(* Logix 5000 project; controller _GigaDiscovery vendor 1 type 14 code 244 rev 35.11; software revision 35.03; part 22 of 23 *)
(* tags used below, declared in another part *)
   All_Rack_Closed_Mem : BOOL;
   Close_Platform_Autocycle_Pylon : BOOL;
   CycleOver : BOOL;
   Emergencies_CL0 : DINT[8];
   FeedBack_Drives_Contactors : BOOL;
   GateCommand : DINT;
   GateRequest : DINT;
   Gates_Auto_Release : BOOL;   // .. At end of Cycle Open Gates Open RESTRAINTS
   Gates_Open_Permissive : Permissive;
   Gondola_Standstill_from_inertia : BOOL;
   HMI_PAGE_PROOF_TEST : DINT;
   I_EStop_Pb_OCC1 : UDT_DCI_STOP_TEST;   // +OCC E-stop -S30301F
   I_EStop_Pb_OCC2 : UDT_DCI_STOP_TEST;   // +OCC2 E-Stop -S28502F
   I_Gondola_Home_Position : BOOL;   // Gondola Home Position -B40002I -B40007I
   I_OCC1_EntGate_PB : BOOL;   // OCC1 Entrance Gate Open/Close -S30701F
   I_OCC1_ExitGate_PB : BOOL;   // OCC1 ExitGate Open/Close -S30707F
   I_OCC2_Disable : UDT_DCM;   // OCC 2 CONTROL DISABLE Page 310
   I_OCC2_ExitGate_PB : BOOL;   // OCC2 ExitGate Open/Close -S28507F
   I_OCC2_RESTRAINTS_RELEASE : Sel_3_Pos_2_Input;   // -S28507F RESTRAINTS RELEASE UNLOCK -RUN- LOCK
   I_OCC_LockOut_Motion : UDT_DCM;   // OCC -Lockout Motion -Q31203E
   I_OCC_Operator_Enable_Key : BOOL;   // OCC Console Enabled -S30305F
   I_Platform_Closed : UDT_DCM;   // Platform Closed RFID Series -B22501J... -B22807J -B22801B
   I_Platform_Line_Min_Pressure_Switch : BOOL;   // Platform Line Minimum Pressure Switch -S21511B
   I_Platform_Line_Unlock_Pressure_Switch : BOOL;   // Unlock Platform Line Pressure Switch -S22006B
   I_Platform_Pressure_on_Close_Circuit : BOOL;   // Platform Maximum Closing Pressure -S21510B
   I_RESTRAINTS_Selector : Sel_3_Pos_2_Input;   // RESTRAINTS Selctor -S30505F Left = Open Right = Close Center = Nothing
   Mem_RESTRAINTS_closed_Correctly : BOOL;
   No_Sfty : Std_to_Sfty;
   O_Close_Gate1 : BOOL;   // Gate 1 OCC2 Operator Close = Mag ON
   O_Close_Gate2 : BOOL;   // Gate 2 Exit Close = Mag ON
   O_Close_Gate3 : BOOL;   // Gate 3 Entrance Close = Mag ON
   O_Close_Gates : BOOL;
   O_Close_Platform : BOOL;
   O_Open_Platform : BOOL;
   O_Platform_Main_Valve : BOOL;   // Valvola principale piattaforma B21902I
   O_RESTRAINTS_MainValve : UDT_CROUT;   // Main Valve -B40501I
   O_RESTRAINTS_Valve_Lift : BOOL;   // Steps 03 04 05
   OS_Start_Stop_Cycle_Started : BOOL;
   Paltform_Cycle_Abborted_Mem : BOOL;   // Paltform Cycle Abborted by Stop Pb Mem
   Pb_Platform_Stop : BOOL;   // Platform Stop Command -S30608F
   PltaformClosed_CycleComplete : BOOL;   // Piattaforme chiuse e ciclo completato
   Power_On_Delay : BOOL;
   ProofTest_Req : BOOL;
   Pylon_Contactor_OFF : BOOL;
   Pylon_Stopped_At_Home : BOOL;   // 5s
   RESTRAINTS_Closed : BOOL;   // All RESTRAINTS Closed
   Restraints_Cycle : Sequencer;
   RESTRAINTS_Left_Press_Switch_Series : BOOL;
   RESTRAINTS_No_Alarms : BOOL;
   Restraints_Permissive : Permissive;
   Restraints_Permissive_Ok : BOOL;
   Restraints_PermissiveLost : DINT;
   RESTRAINTS_Right_Press_Switch_Series : BOOL;
   RESTRAINTS_Sector : LapBars_Sector[9];
   Start_Stop_Cycle : Sequencer;
   Test : DCI_STOP_TEST;
(* S_Platform_and_Gates, continued *)

ROUTINE _10_Gates_Permissive   (* ladder *)
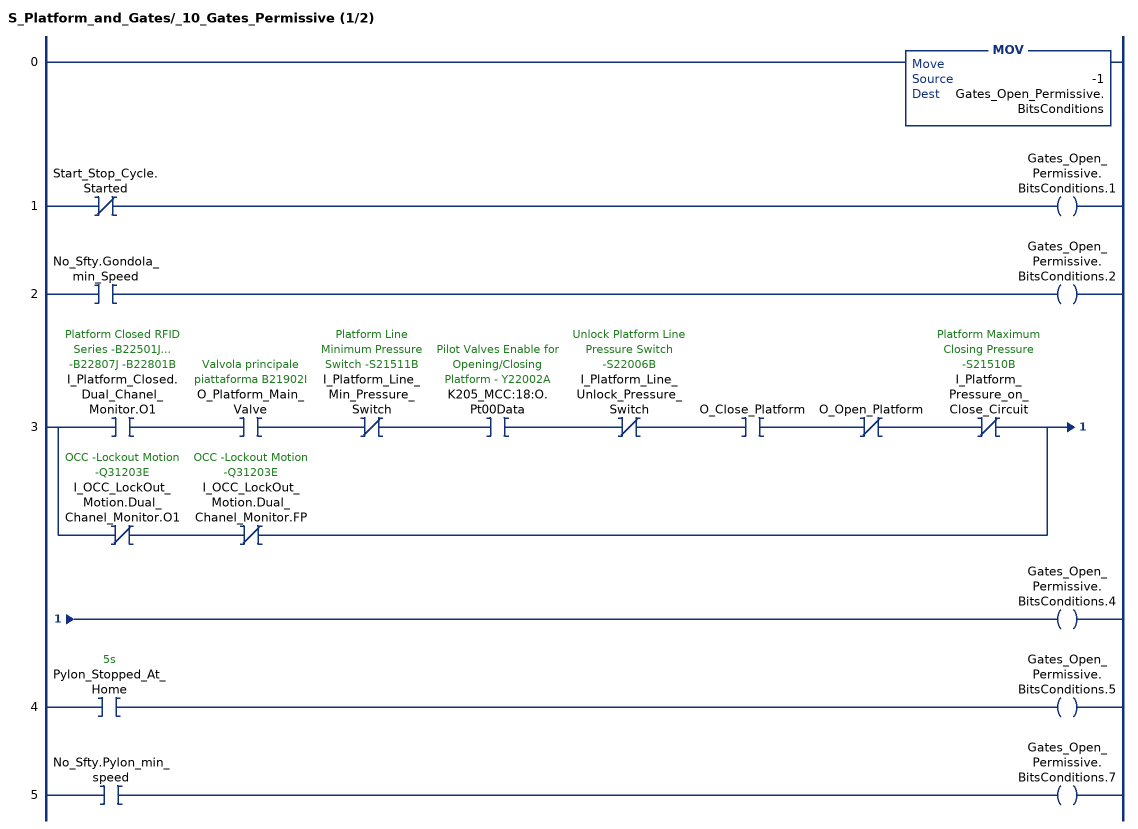
   0: MOV(-1,Gates_Open_Permissive.BitsConditions);
   1: XIO(Start_Stop_Cycle.Started)OTE(Gates_Open_Permissive.BitsConditions.1);
   2: XIC(No_Sfty.Gondola_min_Speed)OTE(Gates_Open_Permissive.BitsConditions.2);
   3: [XIC(I_Platform_Closed.Dual_Chanel_Monitor.O1) XIC(O_Platform_Main_Valve) XIO(I_Platform_Line_Min_Pressure_Switch) XIC(K205_MCC:18:O.Pt00Data) XIO(I_Platform_Line_Unlock_Pressure_Switch) XIC(O_Close_Platform) XIO(O_Open_Platform) XIO(I_Platform_Pressure_on_Close_Circuit) ,XIO(I_OCC_LockOut_Motion.Dual_Chanel_Monitor.O1) XIO(I_OCC_LockOut_Motion.Dual_Chanel_Monitor.FP) ]OTE(Gates_Open_Permissive.BitsConditions.4);
   4: XIC(Pylon_Stopped_At_Home)OTE(Gates_Open_Permissive.BitsConditions.5);
   5: XIC(No_Sfty.Pylon_min_speed)OTE(Gates_Open_Permissive.BitsConditions.7);
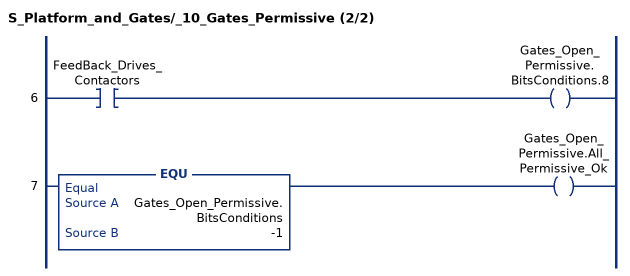
   6: XIC(FeedBack_Drives_Contactors)OTE(Gates_Open_Permissive.BitsConditions.8);
   7: EQU(Gates_Open_Permissive.BitsConditions,-1)OTE(Gates_Open_Permissive.All_Permissive_Ok);
END_ROUTINE

ROUTINE _11_Gates_Commands   (* ladder *)
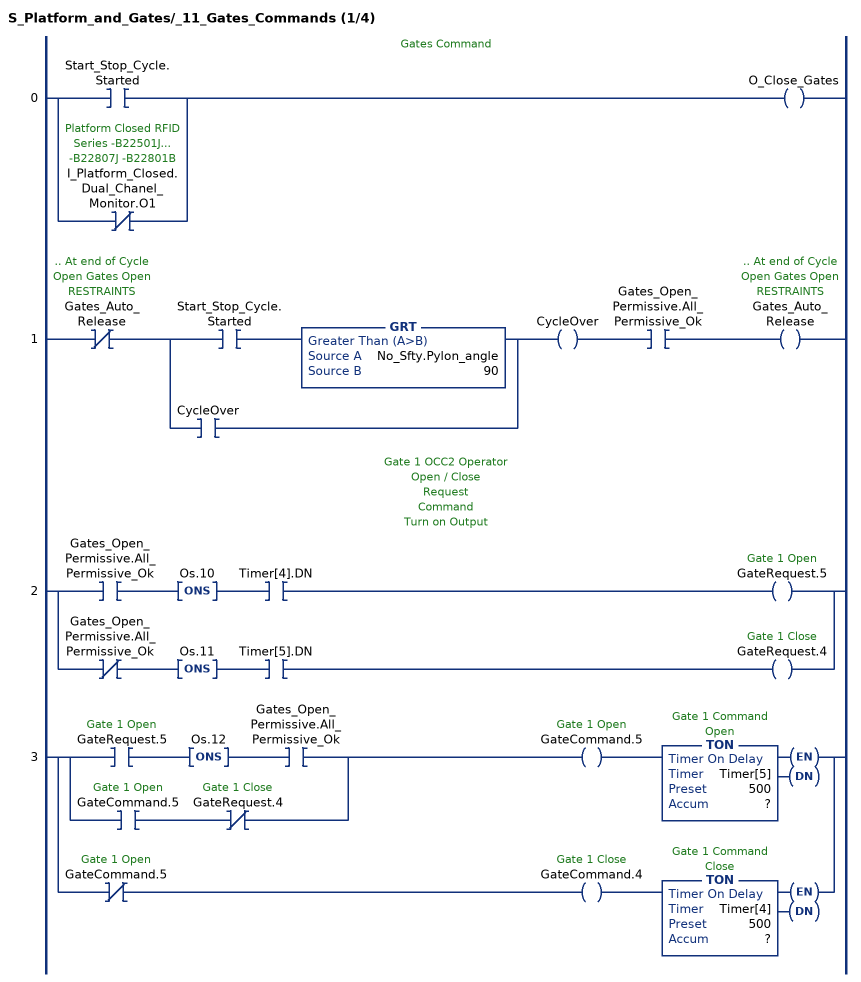
   // Gates Command
   0: [XIC(Start_Stop_Cycle.Started) ,XIO(I_Platform_Closed.Dual_Chanel_Monitor.O1) ]OTE(O_Close_Gates);
   1: XIO(Gates_Auto_Release)[XIC(Start_Stop_Cycle.Started) GRT(No_Sfty.Pylon_angle,90) ,XIC(CycleOver) ]OTE(CycleOver)XIC(Gates_Open_Permissive.All_Permissive_Ok)OTE(Gates_Auto_Release);
   // Gate 1 OCC2 Operator
   // Open / Close
   // Request
   // Command
   // Turn on Output
   2: [XIC(Gates_Open_Permissive.All_Permissive_Ok) ONS(Os.10) XIC(Timer[4].DN) OTE(GateRequest.5) ,XIO(Gates_Open_Permissive.All_Permissive_Ok) ONS(Os.11) XIC(Timer[5].DN) OTE(GateRequest.4) ];
   3: [[XIC(GateRequest.5) ONS(Os.12) XIC(Gates_Open_Permissive.All_Permissive_Ok) ,XIC(GateCommand.5) XIO(GateRequest.4) ] OTE(GateCommand.5) TON(Timer[5],?,?) ,XIO(GateCommand.5) OTE(GateCommand.4) TON(Timer[4],?,?) ];
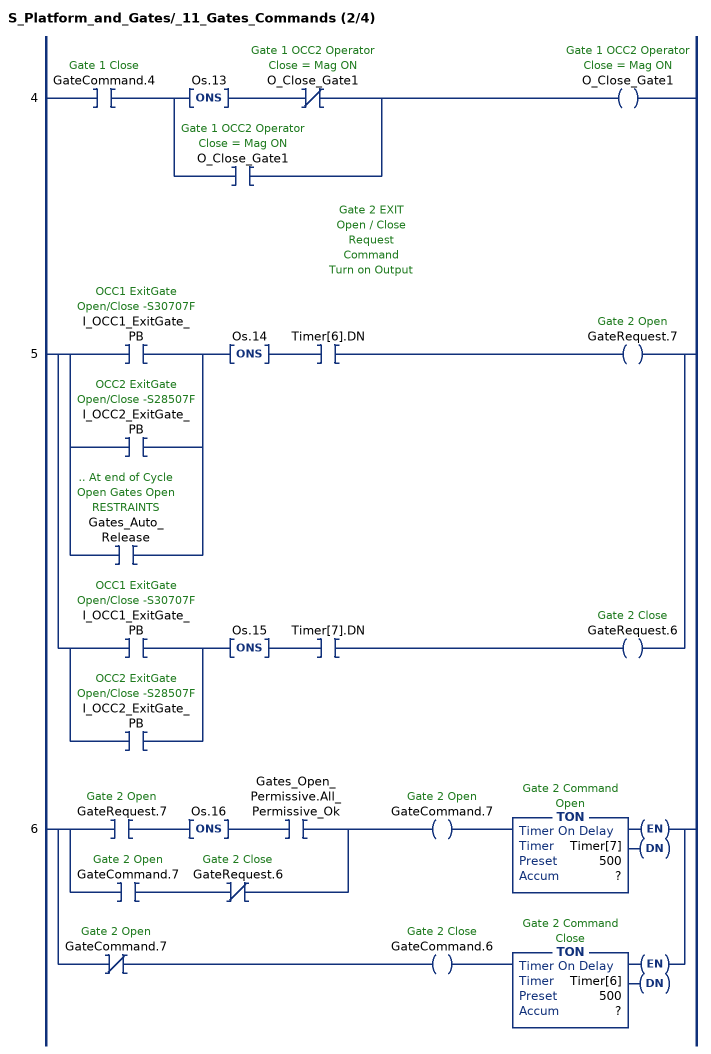
   4: XIC(GateCommand.4)[ONS(Os.13) XIO(O_Close_Gate1) ,XIC(O_Close_Gate1) ]OTE(O_Close_Gate1);
   // Gate 2 EXIT
   // Open / Close
   // Request
   // Command
   // Turn on Output
   5: [[XIC(I_OCC1_ExitGate_PB) ,XIC(I_OCC2_ExitGate_PB) ,XIC(Gates_Auto_Release) ] ONS(Os.14) XIC(Timer[6].DN) OTE(GateRequest.7) ,[XIC(I_OCC1_ExitGate_PB) ,XIC(I_OCC2_ExitGate_PB) ] ONS(Os.15) XIC(Timer[7].DN) OTE(GateRequest.6) ];
   6: [[XIC(GateRequest.7) ONS(Os.16) XIC(Gates_Open_Permissive.All_Permissive_Ok) ,XIC(GateCommand.7) XIO(GateRequest.6) ] OTE(GateCommand.7) TON(Timer[7],?,?) ,XIO(GateCommand.7) OTE(GateCommand.6) TON(Timer[6],?,?) ];
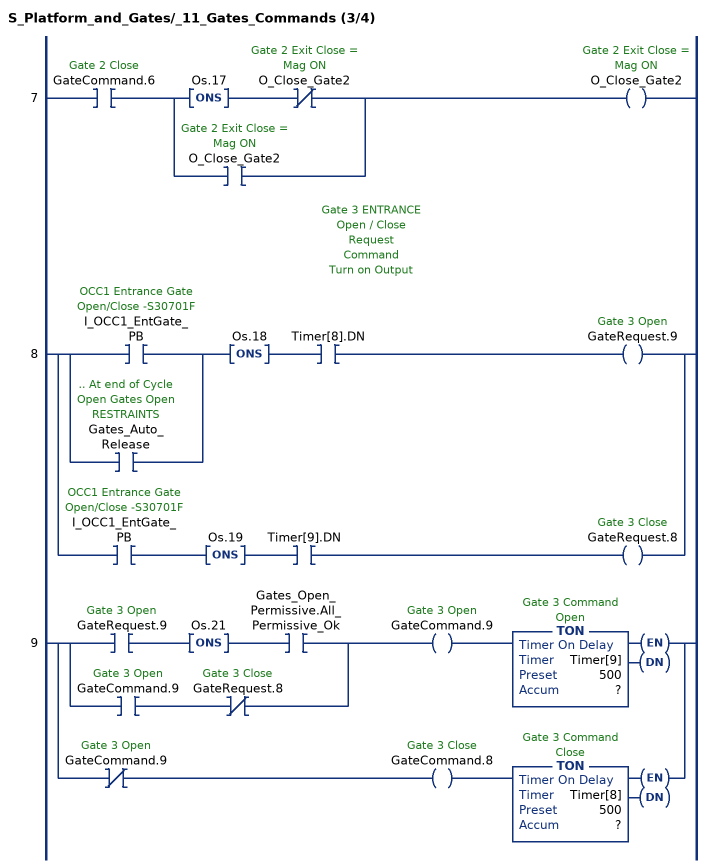
   7: XIC(GateCommand.6)[ONS(Os.17) XIO(O_Close_Gate2) ,XIC(O_Close_Gate2) ]OTE(O_Close_Gate2);
   // Gate 3 ENTRANCE
   // Open / Close
   // Request
   // Command
   // Turn on Output
   8: [[XIC(I_OCC1_EntGate_PB) ,XIC(Gates_Auto_Release) ] ONS(Os.18) XIC(Timer[8].DN) OTE(GateRequest.9) ,XIC(I_OCC1_EntGate_PB) ONS(Os.19) XIC(Timer[9].DN) OTE(GateRequest.8) ];
   9: [[XIC(GateRequest.9) ONS(Os.21) XIC(Gates_Open_Permissive.All_Permissive_Ok) ,XIC(GateCommand.9) XIO(GateRequest.8) ] OTE(GateCommand.9) TON(Timer[9],?,?) ,XIO(GateCommand.9) OTE(GateCommand.8) TON(Timer[8],?,?) ];
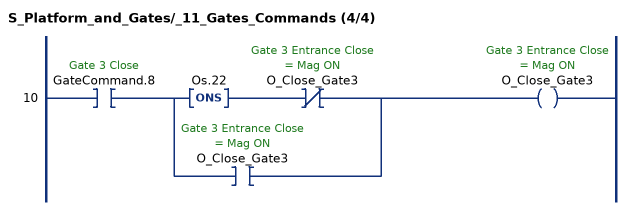
   10: XIC(GateCommand.8)[ONS(Os.22) XIO(O_Close_Gate3) ,XIC(O_Close_Gate3) ]OTE(O_Close_Gate3);
END_ROUTINE

ROUTINE Main   (* ladder *)
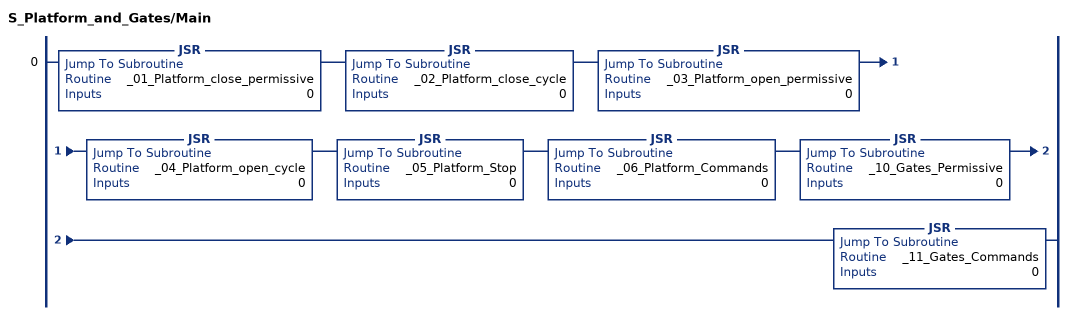
   0: JSR(_01_Platform_close_permissive,0)JSR(_02_Platform_close_cycle,0)JSR(_03_Platform_open_permissive,0)JSR(_04_Platform_open_cycle,0)JSR(_05_Platform_Stop,0)JSR(_06_Platform_Commands,0)JSR(_10_Gates_Permissive,0)JSR(_11_Gates_Commands,0);
END_ROUTINE
END_PROGRAM

PROGRAM S_Restraints_Release   (* main routine Main, safety *)
VAR
   _07_Stop_RESTRAINT_RELEASE_Cycle : BOOL;
   O_Safety_Valve_Unlock_Left_Block : BOOL;   // Steps 02 to 21
   O_Safety_Valve_Unlock_Right_Block : BOOL;   // Steps 02 to 21
   Os : DINT := 45040;
   Proof_Test : Proof_Test := (Validation_Delay_time.PRE := 30000);
   Proof_Test_Req_by_Time : BOOL;
   RESTRAINT_RELEASE_Alarm_Loc : BOOL;
   RESTRAINT_RELEASE_Cycle_AOI : Sequencer_AOI;
   Timer : TIMER[11] := ([0].PRE := 60000, [1].PRE := 2000, [1].ACC := 2000, [1].EN := 1, [1].DN := 1);
END_VAR

ROUTINE _01_Restraints_Release_Permissives   (* ladder *)
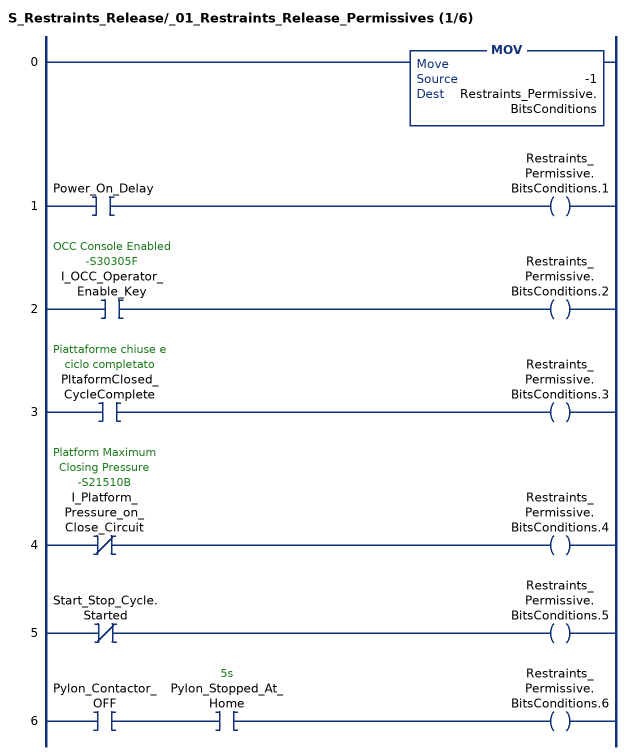
   0: MOV(-1,Restraints_Permissive.BitsConditions);
   1: XIC(Power_On_Delay)OTE(Restraints_Permissive.BitsConditions.1);
   2: XIC(I_OCC_Operator_Enable_Key)OTE(Restraints_Permissive.BitsConditions.2);
   3: XIC(PltaformClosed_CycleComplete)OTE(Restraints_Permissive.BitsConditions.3);
   4: XIO(I_Platform_Pressure_on_Close_Circuit)OTE(Restraints_Permissive.BitsConditions.4);
   5: XIO(Start_Stop_Cycle.Started)OTE(Restraints_Permissive.BitsConditions.5);
   6: XIC(Pylon_Contactor_OFF)XIC(Pylon_Stopped_At_Home)OTE(Restraints_Permissive.BitsConditions.6);
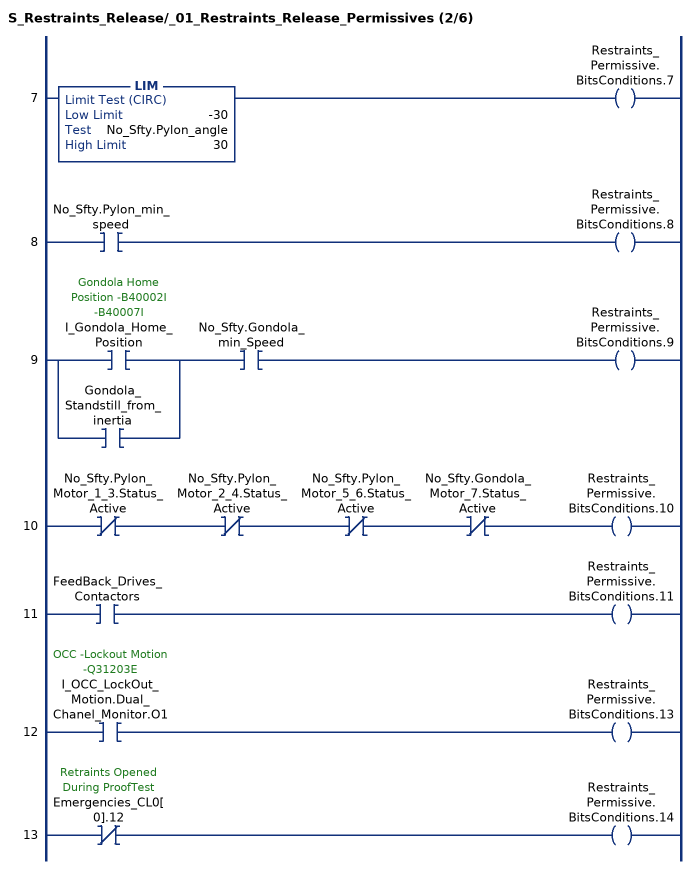
   7: LIM(-30,No_Sfty.Pylon_angle,30)OTE(Restraints_Permissive.BitsConditions.7);
   8: XIC(No_Sfty.Pylon_min_speed)OTE(Restraints_Permissive.BitsConditions.8);
   9: [XIC(I_Gondola_Home_Position) ,XIC(Gondola_Standstill_from_inertia) ]XIC(No_Sfty.Gondola_min_Speed)OTE(Restraints_Permissive.BitsConditions.9);
   10: XIO(No_Sfty.Pylon_Motor_1_3.Status_Active)XIO(No_Sfty.Pylon_Motor_2_4.Status_Active)XIO(No_Sfty.Pylon_Motor_5_6.Status_Active)XIO(No_Sfty.Gondola_Motor_7.Status_Active)OTE(Restraints_Permissive.BitsConditions.10);
   11: XIC(FeedBack_Drives_Contactors)OTE(Restraints_Permissive.BitsConditions.11);
   12: XIC(I_OCC_LockOut_Motion.Dual_Chanel_Monitor.O1)OTE(Restraints_Permissive.BitsConditions.13);
   13: XIO(Emergencies_CL0[0].12)OTE(Restraints_Permissive.BitsConditions.14);
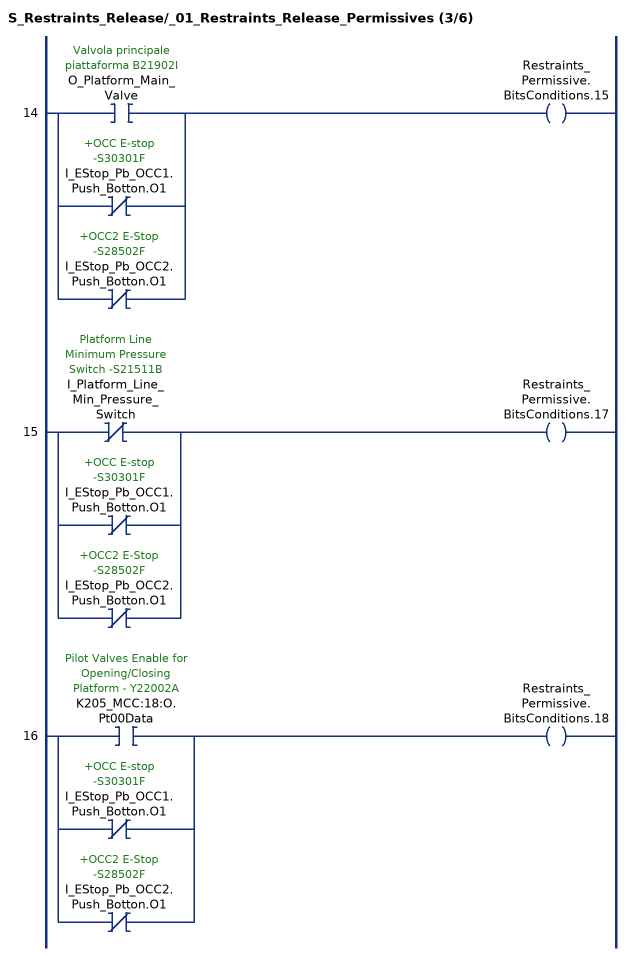
   14: [XIC(O_Platform_Main_Valve) ,XIO(I_EStop_Pb_OCC1.Push_Botton.O1) ,XIO(I_EStop_Pb_OCC2.Push_Botton.O1) ]OTE(Restraints_Permissive.BitsConditions.15);
   15: [XIO(I_Platform_Line_Min_Pressure_Switch) ,XIO(I_EStop_Pb_OCC1.Push_Botton.O1) ,XIO(I_EStop_Pb_OCC2.Push_Botton.O1) ]OTE(Restraints_Permissive.BitsConditions.17);
   16: [XIC(K205_MCC:18:O.Pt00Data) ,XIO(I_EStop_Pb_OCC1.Push_Botton.O1) ,XIO(I_EStop_Pb_OCC2.Push_Botton.O1) ]OTE(Restraints_Permissive.BitsConditions.18);
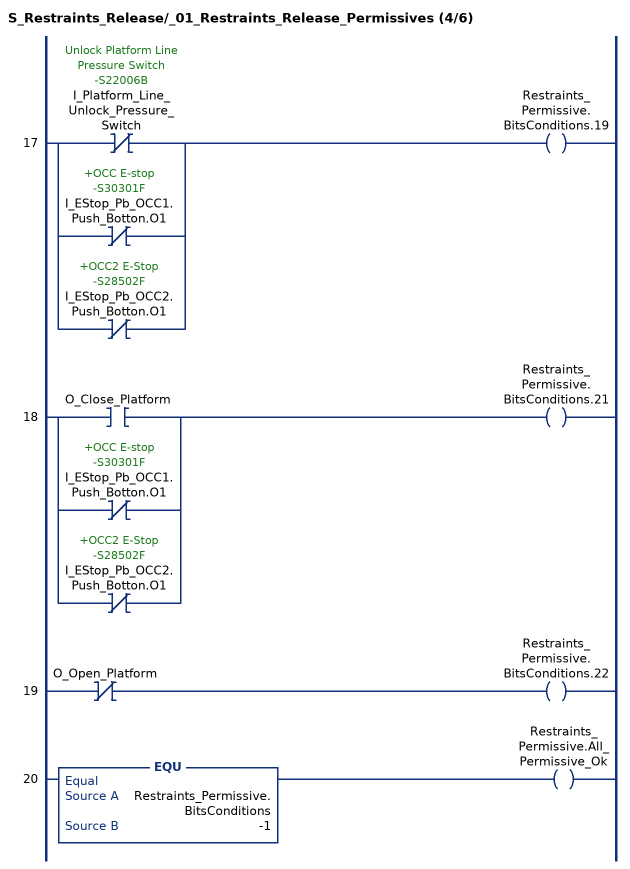
   17: [XIO(I_Platform_Line_Unlock_Pressure_Switch) ,XIO(I_EStop_Pb_OCC1.Push_Botton.O1) ,XIO(I_EStop_Pb_OCC2.Push_Botton.O1) ]OTE(Restraints_Permissive.BitsConditions.19);
   18: [XIC(O_Close_Platform) ,XIO(I_EStop_Pb_OCC1.Push_Botton.O1) ,XIO(I_EStop_Pb_OCC2.Push_Botton.O1) ]OTE(Restraints_Permissive.BitsConditions.21);
   19: XIO(O_Open_Platform)OTE(Restraints_Permissive.BitsConditions.22);
   20: EQU(Restraints_Permissive.BitsConditions,-1)OTE(Restraints_Permissive.All_Permissive_Ok);
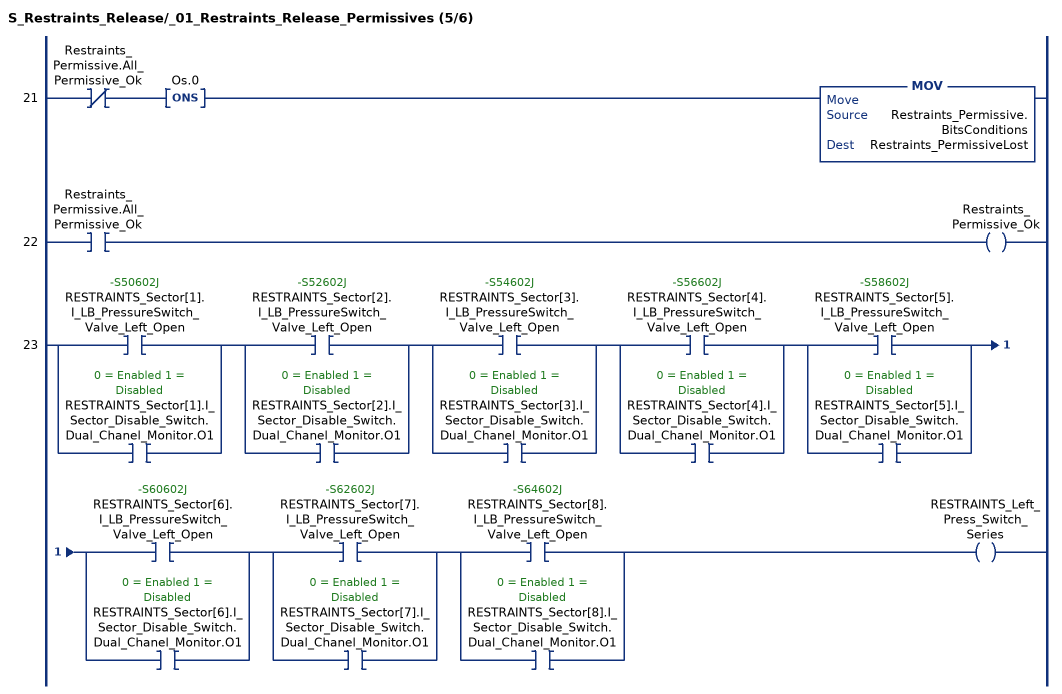
   21: XIO(Restraints_Permissive.All_Permissive_Ok)ONS(Os.0)MOV(Restraints_Permissive.BitsConditions,Restraints_PermissiveLost);
   22: XIC(Restraints_Permissive.All_Permissive_Ok)OTE(Restraints_Permissive_Ok);
   23: [XIC(RESTRAINTS_Sector[1].I_LB_PressureSwitch_Valve_Left_Open) ,XIC(RESTRAINTS_Sector[1].I_Sector_Disable_Switch.Dual_Chanel_Monitor.O1) ][XIC(RESTRAINTS_Sector[2].I_LB_PressureSwitch_Valve_Left_Open) ,XIC(RESTRAINTS_Sector[2].I_Sector_Disable_Switch.Dual_Chanel_Monitor.O1) ][XIC(RESTRAINTS_Sector[3].I_LB_PressureSwitch_Valve_Left_Open) ,XIC(RESTRAINTS_Sector[3].I_Sector_Disable_Switch.Dual_Chanel_Monitor.O1) ][XIC(RESTRAINTS_Sector[4].I_LB_PressureSwitch_Valve_Left_Open) ,XIC(RESTRAINTS_Sector[4].I_Sector_Disable_Switch.Dual_Chanel_Monitor.O1) ][XIC(RESTRAINTS_Sector[5].I_LB_PressureSwitch_Valve_Left_Open) ,XIC(RESTRAINTS_Sector[5].I_Sector_Disable_Switch.Dual_Chanel_Monitor.O1) ][XIC(RESTRAINTS_Sector[6].I_LB_PressureSwitch_Valve_Left_Open) ,XIC(RESTRAINTS_Sector[6].I_Sector_Disable_Switch.Dual_Chanel_Monitor.O1) ][XIC(RESTRAINTS_Sector[7].I_LB_PressureSwitch_Valve_Left_Open) ,XIC(RESTRAINTS_Sector[7].I_Sector_Disable_Switch.Dual_Chanel_Monitor.O1) ][XIC(RESTRAINTS_Sector[8].I_LB_PressureSwitch_Valve_Left_Open) ,XIC(RESTRAINTS_Sector[8].I_Sector_Disable_Switch.Dual_Chanel_Monitor.O1) ]OTE(RESTRAINTS_Left_Press_Switch_Series);
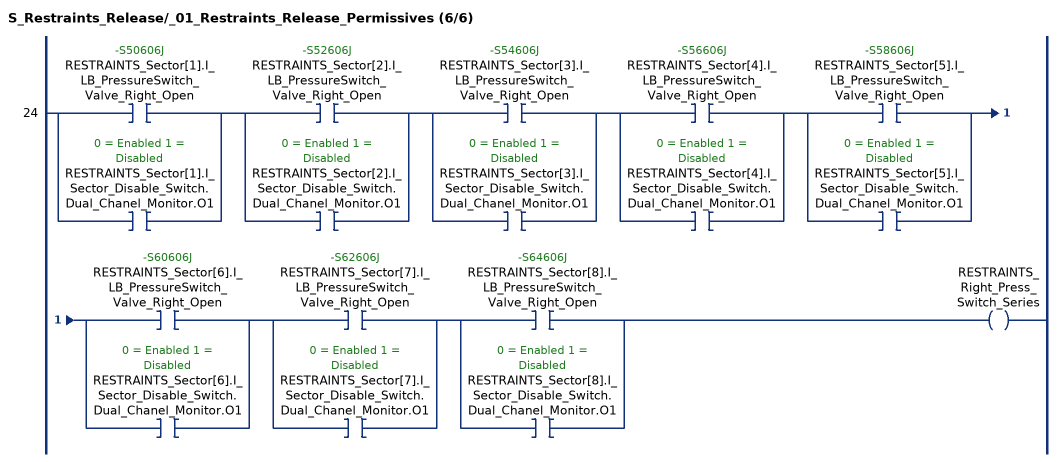
   24: [XIC(RESTRAINTS_Sector[1].I_LB_PressureSwitch_Valve_Right_Open) ,XIC(RESTRAINTS_Sector[1].I_Sector_Disable_Switch.Dual_Chanel_Monitor.O1) ][XIC(RESTRAINTS_Sector[2].I_LB_PressureSwitch_Valve_Right_Open) ,XIC(RESTRAINTS_Sector[2].I_Sector_Disable_Switch.Dual_Chanel_Monitor.O1) ][XIC(RESTRAINTS_Sector[3].I_LB_PressureSwitch_Valve_Right_Open) ,XIC(RESTRAINTS_Sector[3].I_Sector_Disable_Switch.Dual_Chanel_Monitor.O1) ][XIC(RESTRAINTS_Sector[4].I_LB_PressureSwitch_Valve_Right_Open) ,XIC(RESTRAINTS_Sector[4].I_Sector_Disable_Switch.Dual_Chanel_Monitor.O1) ][XIC(RESTRAINTS_Sector[5].I_LB_PressureSwitch_Valve_Right_Open) ,XIC(RESTRAINTS_Sector[5].I_Sector_Disable_Switch.Dual_Chanel_Monitor.O1) ][XIC(RESTRAINTS_Sector[6].I_LB_PressureSwitch_Valve_Right_Open) ,XIC(RESTRAINTS_Sector[6].I_Sector_Disable_Switch.Dual_Chanel_Monitor.O1) ][XIC(RESTRAINTS_Sector[7].I_LB_PressureSwitch_Valve_Right_Open) ,XIC(RESTRAINTS_Sector[7].I_Sector_Disable_Switch.Dual_Chanel_Monitor.O1) ][XIC(RESTRAINTS_Sector[8].I_LB_PressureSwitch_Valve_Right_Open) ,XIC(RESTRAINTS_Sector[8].I_Sector_Disable_Switch.Dual_Chanel_Monitor.O1) ]OTE(RESTRAINTS_Right_Press_Switch_Series);
END_ROUTINE

ROUTINE _02_Restraints_Release_Cycle   (* ladder *)
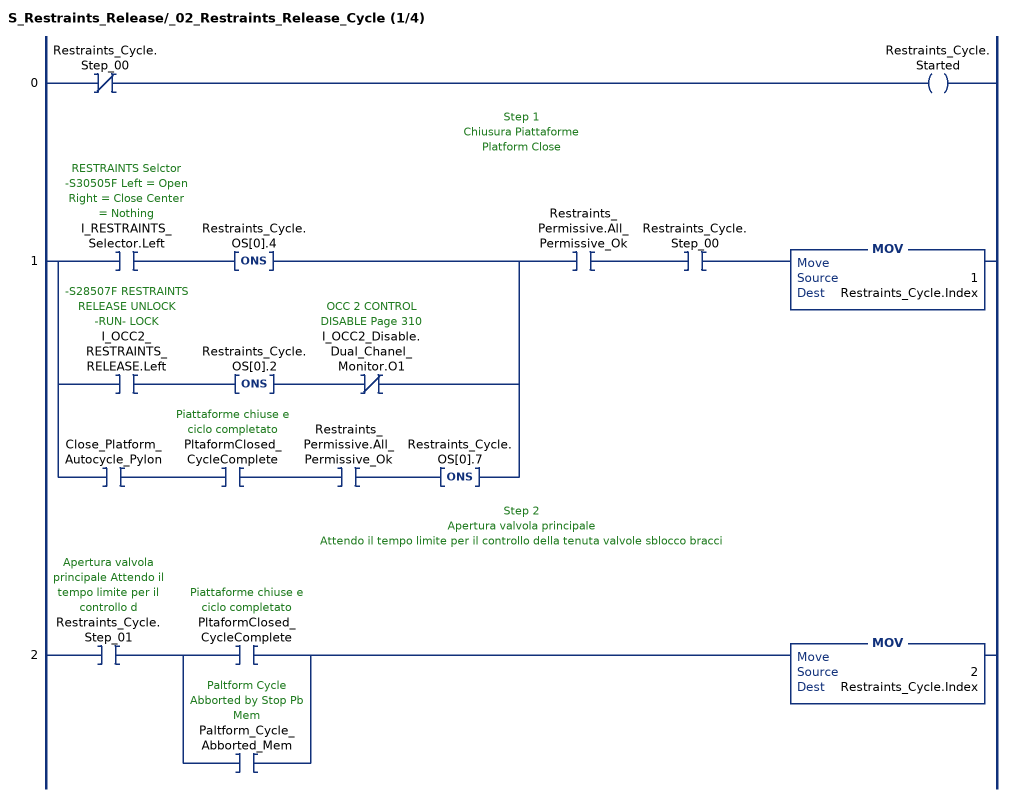
   0: XIO(Restraints_Cycle.Step_00)OTE(Restraints_Cycle.Started);
   // Step 1
   // Chiusura Piattaforme
   // Platform Close
   1: [XIC(I_RESTRAINTS_Selector.Left) ONS(Restraints_Cycle.OS[0].4) ,XIC(I_OCC2_RESTRAINTS_RELEASE.Left) ONS(Restraints_Cycle.OS[0].2) XIO(I_OCC2_Disable.Dual_Chanel_Monitor.O1) ,XIC(Close_Platform_Autocycle_Pylon) XIC(PltaformClosed_CycleComplete) XIC(Restraints_Permissive.All_Permissive_Ok) ONS(Restraints_Cycle.OS[0].7) ]XIC(Restraints_Permissive.All_Permissive_Ok)XIC(Restraints_Cycle.Step_00)MOV(1,Restraints_Cycle.Index);
   // Step 2
   // Apertura valvola principale
   // Attendo il tempo limite per il controllo della tenuta valvole sblocco bracci
   2: XIC(Restraints_Cycle.Step_01)[XIC(PltaformClosed_CycleComplete) ,XIC(Paltform_Cycle_Abborted_Mem) ]MOV(2,Restraints_Cycle.Index);
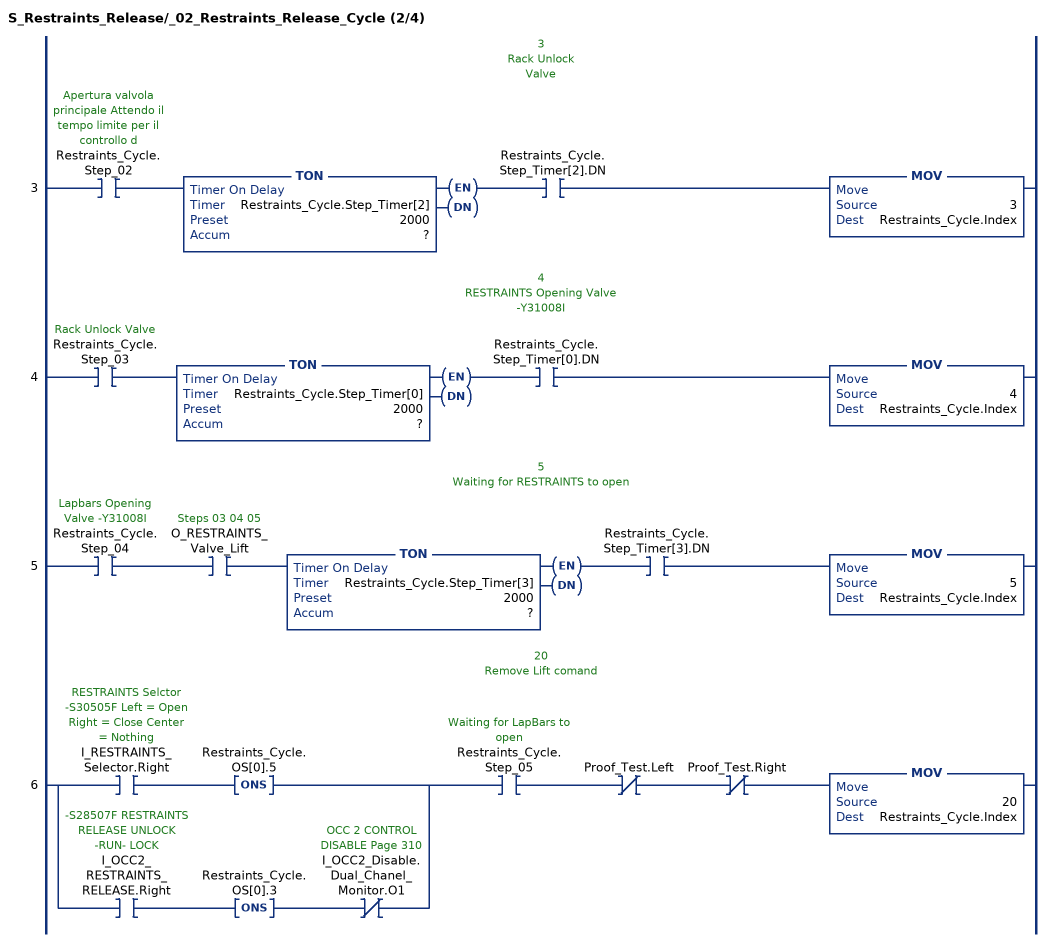
   // 3
   // Rack Unlock
   // Valve
   3: XIC(Restraints_Cycle.Step_02)TON(Restraints_Cycle.Step_Timer[2],?,?)XIC(Restraints_Cycle.Step_Timer[2].DN)MOV(3,Restraints_Cycle.Index);
   // 4
   // RESTRAINTS Opening Valve
   // -Y31008I
   4: XIC(Restraints_Cycle.Step_03)TON(Restraints_Cycle.Step_Timer[0],?,?)XIC(Restraints_Cycle.Step_Timer[0].DN)MOV(4,Restraints_Cycle.Index);
   // 5
   // Waiting for RESTRAINTS to open
   5: XIC(Restraints_Cycle.Step_04)XIC(O_RESTRAINTS_Valve_Lift)TON(Restraints_Cycle.Step_Timer[3],?,?)XIC(Restraints_Cycle.Step_Timer[3].DN)MOV(5,Restraints_Cycle.Index);
   // 20
   // Remove Lift comand
   6: [XIC(I_RESTRAINTS_Selector.Right) ONS(Restraints_Cycle.OS[0].5) ,XIC(I_OCC2_RESTRAINTS_RELEASE.Right) ONS(Restraints_Cycle.OS[0].3) XIO(I_OCC2_Disable.Dual_Chanel_Monitor.O1) ]XIC(Restraints_Cycle.Step_05)XIO(Proof_Test.Left)XIO(Proof_Test.Right)MOV(20,Restraints_Cycle.Index);
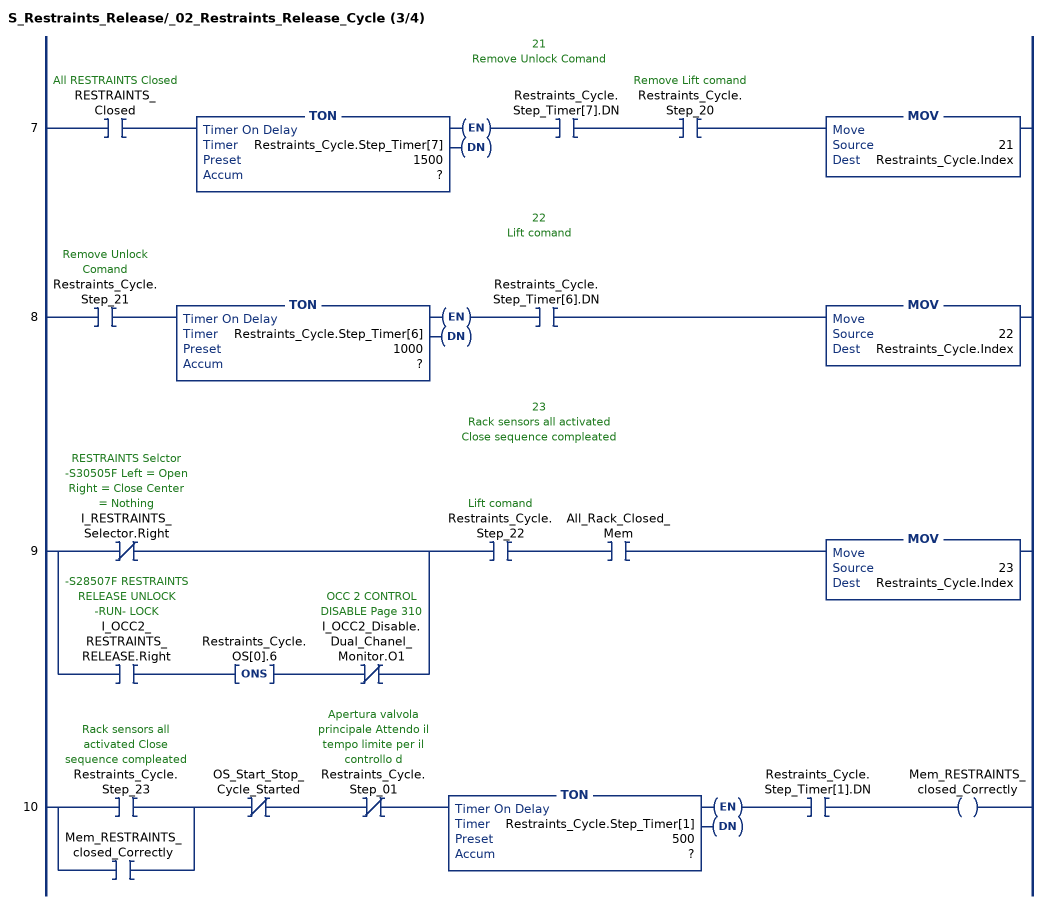
   // 21
   // Remove Unlock Comand
   7: XIC(RESTRAINTS_Closed)TON(Restraints_Cycle.Step_Timer[7],?,?)XIC(Restraints_Cycle.Step_Timer[7].DN)XIC(Restraints_Cycle.Step_20)MOV(21,Restraints_Cycle.Index);
   // 22
   // Lift comand
   8: XIC(Restraints_Cycle.Step_21)TON(Restraints_Cycle.Step_Timer[6],?,?)XIC(Restraints_Cycle.Step_Timer[6].DN)MOV(22,Restraints_Cycle.Index);
   // 23
   // Rack sensors all activated
   // Close sequence compleated
   9: [XIO(I_RESTRAINTS_Selector.Right) ,XIC(I_OCC2_RESTRAINTS_RELEASE.Right) ONS(Restraints_Cycle.OS[0].6) XIO(I_OCC2_Disable.Dual_Chanel_Monitor.O1) ]XIC(Restraints_Cycle.Step_22)XIC(All_Rack_Closed_Mem)MOV(23,Restraints_Cycle.Index);
   10: [XIC(Restraints_Cycle.Step_23) ,XIC(Mem_RESTRAINTS_closed_Correctly) ]XIO(OS_Start_Stop_Cycle_Started)XIO(Restraints_Cycle.Step_01)TON(Restraints_Cycle.Step_Timer[1],?,?)XIC(Restraints_Cycle.Step_Timer[1].DN)OTE(Mem_RESTRAINTS_closed_Correctly);
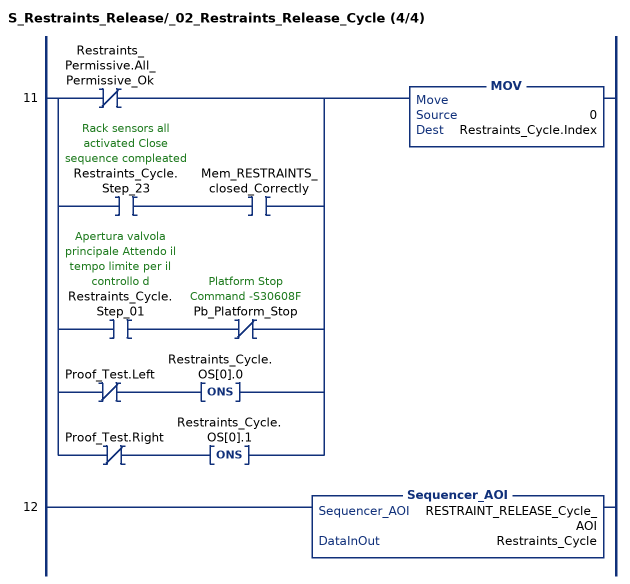
   11: [XIO(Restraints_Permissive.All_Permissive_Ok) ,XIC(Restraints_Cycle.Step_23) XIC(Mem_RESTRAINTS_closed_Correctly) ,XIC(Restraints_Cycle.Step_01) XIO(Pb_Platform_Stop) ,XIO(Proof_Test.Left) ONS(Restraints_Cycle.OS[0].0) ,XIO(Proof_Test.Right) ONS(Restraints_Cycle.OS[0].1) ]MOV(0,Restraints_Cycle.Index);
   12: Sequencer_AOI(RESTRAINT_RELEASE_Cycle_AOI,Restraints_Cycle);
END_ROUTINE

ROUTINE _03_Proof_Test   (* ladder *)
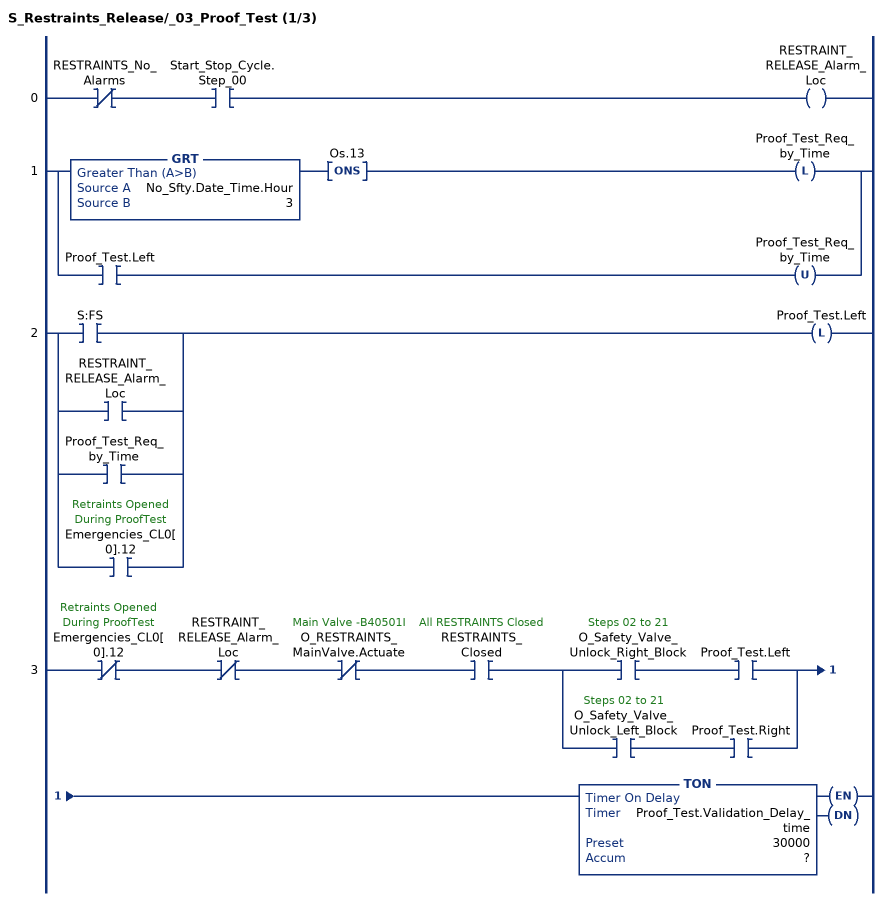
   0: XIO(RESTRAINTS_No_Alarms)XIC(Start_Stop_Cycle.Step_00)OTE(RESTRAINT_RELEASE_Alarm_Loc);
   1: [GRT(No_Sfty.Date_Time.Hour,3) ONS(Os.13) OTL(Proof_Test_Req_by_Time) ,XIC(Proof_Test.Left) OTU(Proof_Test_Req_by_Time) ];
   2: [XIC(S:FS) ,XIC(RESTRAINT_RELEASE_Alarm_Loc) ,XIC(Proof_Test_Req_by_Time) ,XIC(Emergencies_CL0[0].12) ]OTL(Proof_Test.Left);
   3: XIO(Emergencies_CL0[0].12)XIO(RESTRAINT_RELEASE_Alarm_Loc)XIO(O_RESTRAINTS_MainValve.Actuate)XIC(RESTRAINTS_Closed)[XIC(O_Safety_Valve_Unlock_Right_Block) XIC(Proof_Test.Left) ,XIC(O_Safety_Valve_Unlock_Left_Block) XIC(Proof_Test.Right) ]TON(Proof_Test.Validation_Delay_time,?,?);
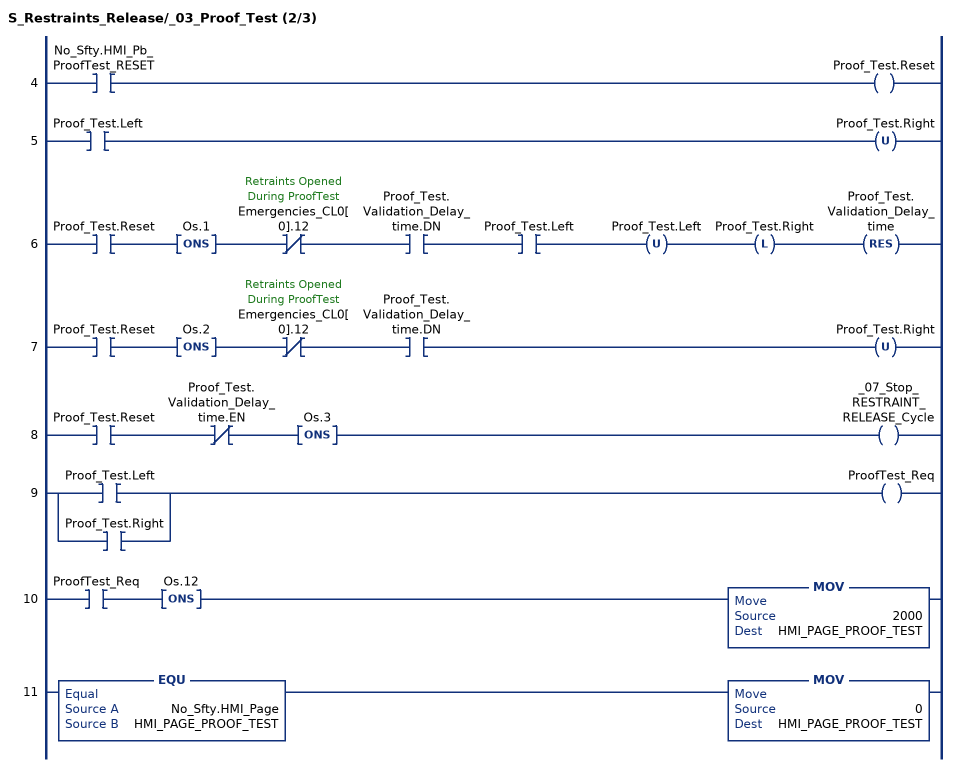
   4: XIC(No_Sfty.HMI_Pb_ProofTest_RESET)OTE(Proof_Test.Reset);
   5: XIC(Proof_Test.Left)OTU(Proof_Test.Right);
   6: XIC(Proof_Test.Reset)ONS(Os.1)XIO(Emergencies_CL0[0].12)XIC(Proof_Test.Validation_Delay_time.DN)XIC(Proof_Test.Left)OTU(Proof_Test.Left)OTL(Proof_Test.Right)RES(Proof_Test.Validation_Delay_time);
   7: XIC(Proof_Test.Reset)ONS(Os.2)XIO(Emergencies_CL0[0].12)XIC(Proof_Test.Validation_Delay_time.DN)OTU(Proof_Test.Right);
   8: XIC(Proof_Test.Reset)XIO(Proof_Test.Validation_Delay_time.EN)ONS(Os.3)OTE(_07_Stop_RESTRAINT_RELEASE_Cycle);
   9: [XIC(Proof_Test.Left) ,XIC(Proof_Test.Right) ]OTE(ProofTest_Req);
   10: XIC(ProofTest_Req)ONS(Os.12)MOV(2000,HMI_PAGE_PROOF_TEST);
   11: EQU(No_Sfty.HMI_Page,HMI_PAGE_PROOF_TEST)MOV(0,HMI_PAGE_PROOF_TEST);
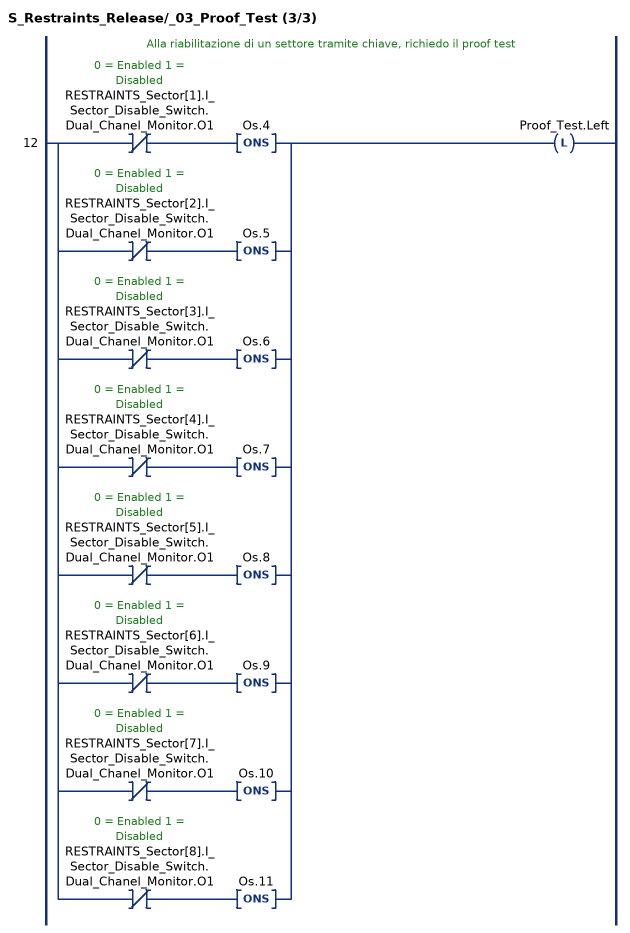
   // Alla riabilitazione di un settore tramite chiave, richiedo il proof test
   12: [XIO(RESTRAINTS_Sector[1].I_Sector_Disable_Switch.Dual_Chanel_Monitor.O1) ONS(Os.4) ,XIO(RESTRAINTS_Sector[2].I_Sector_Disable_Switch.Dual_Chanel_Monitor.O1) ONS(Os.5) ,XIO(RESTRAINTS_Sector[3].I_Sector_Disable_Switch.Dual_Chanel_Monitor.O1) ONS(Os.6) ,XIO(RESTRAINTS_Sector[4].I_Sector_Disable_Switch.Dual_Chanel_Monitor.O1) ONS(Os.7) ,XIO(RESTRAINTS_Sector[5].I_Sector_Disable_Switch.Dual_Chanel_Monitor.O1) ONS(Os.8) ,XIO(RESTRAINTS_Sector[6].I_Sector_Disable_Switch.Dual_Chanel_Monitor.O1) ONS(Os.9) ,XIO(RESTRAINTS_Sector[7].I_Sector_Disable_Switch.Dual_Chanel_Monitor.O1) ONS(Os.10) ,XIO(RESTRAINTS_Sector[8].I_Sector_Disable_Switch.Dual_Chanel_Monitor.O1) ONS(Os.11) ]OTL(Proof_Test.Left);
END_ROUTINE
